   "Carrier_81_G120DStatusWord.9" AT %I4413.1 : Bool;   // Bit_09_CONTR_PLC
   "Carrier_81_G120DStatusWord.10" AT %I4413.2 : Bool;   // Bit_10_F_MAX
   "Carrier_81_G120DStatusWord.11" AT %I4413.3 : Bool;   // Bit_11_LIMIT_REACHED
   "Carrier_81_G120DStatusWord.12" AT %I4413.4 : Bool;   // Bit_12_BRAKE_OPEN
   "Carrier_81_G120DStatusWord.13" AT %I4413.5 : Bool;   // Bit_13_NO_OVERTEMP
   "Carrier_81_G120DStatusWord.14" AT %I4413.6 : Bool;   // Bit_14_CW_CCW
   "Carrier_81_G120DStatusWord.15" AT %I4413.7 : Bool;   // Bit_15_OVERL
   "Carrier_81_Slot2_Input" AT %IW4414 : Word;   // SLOT 2 INPUT WORD
   "Carrier_81_CrashDetectSW" AT %I4414.0 : Bool;   // CRASH DETECT SW
   "Carrier_81_SpareSafetyInput(2_1)" AT %I4414.1 : Bool;   // SPARE SAFETY INPUT
   "Carrier_81_SpareSafetyInput(2_2)" AT %I4414.2 : Bool;   // SPARE SAFETY INPUT
   "Carrier_81_SpareSafetyInput(2_3)" AT %I4414.3 : Bool;   // SPARE SAFETY INPUT
   "Carrier_81_SpareSafetyInput(2_4)" AT %I4414.4 : Bool;   // SPARE SAFETY INPUT
   "Carrier_81_SpareSafetyInput(2_5)" AT %I4414.5 : Bool;   // SPARE SAFETY INPUT
   "Carrier_81_SpareSafetyInput(2_6)" AT %I4414.6 : Bool;   // SPARE SAFETY INPUT
   "Carrier_81_SpareSafetyInput(2_7)" AT %I4414.7 : Bool;   // SPARE SAFETY INPUT
   "Carrier_81_Slot3_SafetyOutput" AT %IW4415 : Word;   // SLOT 3 SAFETY OUTPUT WORD
   "Carrier_81_Crash_Detect_OK" AT %I4415.0 : Bool;   // CARRIER CRASH DETECT
   "Carrier_81_SpareSafetyOutput(3_1)" AT %I4415.1 : Bool;   // SPARE SAFETY OUTPUT
   "Carrier_81_SpareSafetyOutput(3_2)" AT %I4415.2 : Bool;   // SPARE SAFETY OUTPUT
   "Carrier_81_SpareSafetyOutput(3_3)" AT %I4415.3 : Bool;   // SPARE SAFETY OUTPUT
   "Carrier_81_SpareSafetyOutput(3_4)" AT %I4415.4 : Bool;   // SPARE SAFETY OUTPUT
   "Carrier_81_SpareSafetyOutput(3_5)" AT %I4415.5 : Bool;   // SPARE SAFETY OUTPUT
   "Carrier_81_SpareSafetyOutput(3_6)" AT %I4415.6 : Bool;   // SPARE SAFETY OUTPUT
   "Carrier_81_SpareSafetyOutput(3_7)" AT %I4415.7 : Bool;   // SPARE SAFETY OUTPUT
   "Carrier_81_Slot4_Input" AT %IW4416 : Word;   // SLOT 4 INPUT WORD
   "Carrier_81_480VPowerOn_MDCB1" AT %I4416.0 : Bool;   // 480 VAC POWER ON MDCB 1
   "Carrier_81_SpareInput(4_1)" AT %I4416.1 : Bool;   // SPARE INPUT
   "Carrier_81_SpareInput(4_2)" AT %I4416.2 : Bool;   // SPARE INPUT
   "Carrier_81_SitopSelectStatus" AT %I4416.3 : Bool;   // SITOP SELECT STATUS
   "Carrier_81_DCsupplyOnPSCB2" AT %I4416.4 : Bool;   // DC SUPPLY ON PSCB 2
   "Carrier_81_SpareInput(4_5)" AT %I4416.5 : Bool;   // SPARE INPUT
   "Carrier_81_SpareInput(4_6)" AT %I4416.6 : Bool;   // SPARE INPUT
   "Carrier_81_SpareInput(4_7)" AT %I4416.7 : Bool;   // SPARE INPUT
   "Carrier_81_PB1_ProdHoldLH" AT %I4417.0 : Bool;   // PB 1 PRODUCTION HOLD LH
   "Carrier_81_PB2_ResetLH" AT %I4417.1 : Bool;   // PB 2 RESET LH
   "Carrier_81_PB3_ProdHoldRH" AT %I4417.2 : Bool;   // PB 3 PRODUCTION HOLD RH
   "Carrier_81_PB4_ResetRH" AT %I4417.3 : Bool;   // PB 4 RESET RH
   "Carrier_81_SpareInput(4_14)" AT %I4417.4 : Bool;   // SPARE INPUT
   "Carrier_81_SpareInput(4_15)" AT %I4417.5 : Bool;   // SPARE INPUT
   "Carrier_81_SpareInput(4_16)" AT %I4417.6 : Bool;   // SPARE INPUT
   "Carrier_81_SpareInput(4_17)" AT %I4417.7 : Bool;   // SPARE INPUT
   "Carrier_81_Slot5_Output" AT %IW4418 : Word;   // SLOT 5 OUTPUT WORD
   "Carrier_81_IRD400_HMI_24VDC_ENABLE" AT %I4418.0 : Bool;   // IRD 400 PANEL HMI 24V DC POWER
   "Carrier_81_FaultLight_LH" AT %I4418.1 : Bool;   // FAULT LIGHT LH
   "Carrier_81_RunLight_LH" AT %I4418.2 : Bool;   // RUN LIGHT LH
   "Carrier_81_FaultLight_RH" AT %I4418.3 : Bool;   // FAULT LIGHT RH
   "Carrier_81_RunLight_RH" AT %I4418.4 : Bool;   // RUN LIGHT RH
   "Carrier_81_SpareOutput(5_5)" AT %I4418.5 : Bool;   // SPARE OUTPUT
   "Carrier_81_SpareOutput(5_6)" AT %I4418.6 : Bool;   // SPARE OUTPUT
   "Carrier_81_SpareOutput(5_7)" AT %I4418.7 : Bool;   // SPARE OUTPUT
   "Carrier_81_ActualSpeed" AT %IW4420 : Word;   // ACTUAL SPEED
   "Carrier_81_CarrierDriveAlarm" AT %IW4422 : Word;   // CARRIER DRIVE ALARM
   "Carrier_81_CarrierDriveWarning" AT %IW4424 : Word;   // CARRIER DRIVE WARNING
   "Carrier_82_Status" AT %IW4450 : Word;   // CARRIER STATUS WORD
   "Carrier_82_Status.0" AT %I4450.0 : Bool;   // HEARTBEAT
   "Carrier_82_Status.1" AT %I4450.1 : Bool;   // MANUAL
   "Carrier_82_Status.2" AT %I4450.2 : Bool;   // IN_AUTO
   "Carrier_82_Status.3" AT %I4450.3 : Bool;   // POSITIONING_COMPLETE
   "Carrier_82_Status.4" AT %I4450.4 : Bool;   // PRODUCTION HOLD
   "Carrier_82_Status.5" AT %I4450.5 : Bool;   // CARRIER MOVING FORWARD
   "Carrier_82_Status.6" AT %I4450.6 : Bool;   // CARRIER MOVING REVERSE
   "Carrier_82_Status.7" AT %I4450.7 : Bool;   // CARRIER FAULT
   "Carrier_82_Status.8" AT %I4451.0 : Bool;   // CRASH DETECT TRIPPED
   "Carrier_82_Status.9" AT %I4451.1 : Bool;
   "Carrier_82_Status.10" AT %I4451.2 : Bool;
   "Carrier_82_Status.11" AT %I4451.3 : Bool;
   "Carrier_82_Status.12" AT %I4451.4 : Bool;
   "Carrier_82_Status.13" AT %I4451.5 : Bool;
   "Carrier_82_Status.14" AT %I4451.6 : Bool;
   "Carrier_82_Status.15" AT %I4451.7 : Bool;
   "Carrier_82_SDCFaultCode" AT %IW4452 : Word;   // SDC FAULT CODE
   "Carrier_82_CarrierPosition" AT %ID4454 : DWord;   // CARRIER POSITION
   "Carrier_82_CarrierNumber" AT %IW4458 : Word;   // CARRIER NUMBER
   "Carrier_82_G120DControlWord" AT %IW4460 : Word;   // G120D_STW1_CONTROL
   "Carrier_82_G120DControlWord.0" AT %I4460.0 : Bool;   // Bit_00_ON
   "Carrier_82_G120DControlWord.1" AT %I4460.1 : Bool;   // Bit_01_AUS2_INH
   "Carrier_82_G120DControlWord.2" AT %I4460.2 : Bool;   // Bit_02_AUS3_STOP
   "Carrier_82_G120DControlWord.3" AT %I4460.3 : Bool;   // Bit_03_EN
   "Carrier_82_G120DControlWord.4" AT %I4460.4 : Bool;   // Bit_04_EN_RAMP
   "Carrier_82_G120DControlWord.5" AT %I4460.5 : Bool;   // Bit_05_START_RAMP
   "Carrier_82_G120DControlWord.6" AT %I4460.6 : Bool;   // Bit_06_SETPOINT
   "Carrier_82_G120DControlWord.7" AT %I4460.7 : Bool;   // Bit_07_RESET
   "Carrier_82_G120DControlWord.8" AT %I4461.0 : Bool;   // Bit_08_JOG_R
   "Carrier_82_G120DControlWord.9" AT %I4461.1 : Bool;   // Bit_09_JOG_L
   "Carrier_82_G120DControlWord.10" AT %I4461.2 : Bool;   // Bit_10_CONTR_PLC
   "Carrier_82_G120DControlWord.11" AT %I4461.3 : Bool;   // Bit_11_REVERSE
   "Carrier_82_G120DControlWord.12" AT %I4461.4 : Bool;   // Bit_12_BRAKE_RELEASE
   "Carrier_82_G120DControlWord.13" AT %I4461.5 : Bool;   // Bit_13_DDS
   "Carrier_82_G120DControlWord.14" AT %I4461.6 : Bool;   // Bit_14_DO0
   "Carrier_82_G120DControlWord.15" AT %I4461.7 : Bool;   // Bit_15_DO1
   "Carrier_82_G120DStatusWord" AT %IW4462 : Word;   // G120D_ZSW1_STATUS
   "Carrier_82_G120DStatusWord.0" AT %I4462.0 : Bool;   // Bit_00_READY_RUN
   "Carrier_82_G120DStatusWord.1" AT %I4462.1 : Bool;   // Bit_01_READY_ON
   "Carrier_82_G120DStatusWord.2" AT %I4462.2 : Bool;   // Bit_02_ENABLE
   "Carrier_82_G120DStatusWord.3" AT %I4462.3 : Bool;   // Bit_03_FAULT
   "Carrier_82_G120DStatusWord.4" AT %I4462.4 : Bool;   // Bit_04_OFF2
   "Carrier_82_G120DStatusWord.5" AT %I4462.5 : Bool;   // Bit_05_OFF3
   "Carrier_82_G120DStatusWord.6" AT %I4462.6 : Bool;   // Bit_06_LOCK_OUT
   "Carrier_82_G120DStatusWord.7" AT %I4462.7 : Bool;   // Bit_07_WARN
   "Carrier_82_G120DStatusWord.8" AT %I4463.0 : Bool;   // Bit_08_NO_DEVIATION
   "Carrier_82_G120DStatusWord.9" AT %I4463.1 : Bool;   // Bit_09_CONTR_PLC
   "Carrier_82_G120DStatusWord.10" AT %I4463.2 : Bool;   // Bit_10_F_MAX
   "Carrier_82_G120DStatusWord.11" AT %I4463.3 : Bool;   // Bit_11_LIMIT_REACHED
   "Carrier_82_G120DStatusWord.12" AT %I4463.4 : Bool;   // Bit_12_BRAKE_OPEN
   "Carrier_82_G120DStatusWord.13" AT %I4463.5 : Bool;   // Bit_13_NO_OVERTEMP
   "Carrier_82_G120DStatusWord.14" AT %I4463.6 : Bool;   // Bit_14_CW_CCW
   "Carrier_82_G120DStatusWord.15" AT %I4463.7 : Bool;   // Bit_15_OVERL
   "Carrier_82_Slot2_Input" AT %IW4464 : Word;   // SLOT 2 INPUT WORD
   "Carrier_82_CrashDetectSW" AT %I4464.0 : Bool;   // CRASH DETECT SW
   "Carrier_82_SpareSafetyInput(2_1)" AT %I4464.1 : Bool;   // SPARE SAFETY INPUT
   "Carrier_82_SpareSafetyInput(2_2)" AT %I4464.2 : Bool;   // SPARE SAFETY INPUT
   "Carrier_82_SpareSafetyInput(2_3)" AT %I4464.3 : Bool;   // SPARE SAFETY INPUT
   "Carrier_82_SpareSafetyInput(2_4)" AT %I4464.4 : Bool;   // SPARE SAFETY INPUT
   "Carrier_82_SpareSafetyInput(2_5)" AT %I4464.5 : Bool;   // SPARE SAFETY INPUT
   "Carrier_82_SpareSafetyInput(2_6)" AT %I4464.6 : Bool;   // SPARE SAFETY INPUT
   "Carrier_82_SpareSafetyInput(2_7)" AT %I4464.7 : Bool;   // SPARE SAFETY INPUT
   "Carrier_82_Slot3_SafetyOutput" AT %IW4465 : Word;   // SLOT 3 SAFETY OUTPUT WORD
   "Carrier_82_Crash_Detect_OK" AT %I4465.0 : Bool;   // CARRIER CRASH DETECT
   "Carrier_82_SpareSafetyOutput(3_1)" AT %I4465.1 : Bool;   // SPARE SAFETY OUTPUT
   "Carrier_82_SpareSafetyOutput(3_2)" AT %I4465.2 : Bool;   // SPARE SAFETY OUTPUT
   "Carrier_82_SpareSafetyOutput(3_3)" AT %I4465.3 : Bool;   // SPARE SAFETY OUTPUT
   "Carrier_82_SpareSafetyOutput(3_4)" AT %I4465.4 : Bool;   // SPARE SAFETY OUTPUT
   "Carrier_82_SpareSafetyOutput(3_5)" AT %I4465.5 : Bool;   // SPARE SAFETY OUTPUT
   "Carrier_82_SpareSafetyOutput(3_6)" AT %I4465.6 : Bool;   // SPARE SAFETY OUTPUT
   "Carrier_82_SpareSafetyOutput(3_7)" AT %I4465.7 : Bool;   // SPARE SAFETY OUTPUT
   "Carrier_82_Slot4_Input" AT %IW4466 : Word;   // SLOT 4 INPUT WORD
   "Carrier_82_480VPowerOn_MDCB1" AT %I4466.0 : Bool;   // 480 VAC POWER ON MDCB 1
   "Carrier_82_SpareInput(4_1)" AT %I4466.1 : Bool;   // SPARE INPUT
   "Carrier_82_SpareInput(4_2)" AT %I4466.2 : Bool;   // SPARE INPUT
   "Carrier_82_SitopSelectStatus" AT %I4466.3 : Bool;   // SITOP SELECT STATUS
   "Carrier_82_DCsupplyOnPSCB2" AT %I4466.4 : Bool;   // DC SUPPLY ON PSCB 2
   "Carrier_82_SpareInput(4_5)" AT %I4466.5 : Bool;   // SPARE INPUT
   "Carrier_82_SpareInput(4_6)" AT %I4466.6 : Bool;   // SPARE INPUT
   "Carrier_82_SpareInput(4_7)" AT %I4466.7 : Bool;   // SPARE INPUT
   "Carrier_82_PB1_ProdHoldLH" AT %I4467.0 : Bool;   // PB 1 PRODUCTION HOLD LH
   "Carrier_82_PB2_ResetLH" AT %I4467.1 : Bool;   // PB 2 RESET LH
   "Carrier_82_PB3_ProdHoldRH" AT %I4467.2 : Bool;   // PB 3 PRODUCTION HOLD RH
   "Carrier_82_PB4_ResetRH" AT %I4467.3 : Bool;   // PB 4 RESET RH
   "Carrier_82_SpareInput(4_14)" AT %I4467.4 : Bool;   // SPARE INPUT
   "Carrier_82_SpareInput(4_15)" AT %I4467.5 : Bool;   // SPARE INPUT
   "Carrier_82_SpareInput(4_16)" AT %I4467.6 : Bool;   // SPARE INPUT
   "Carrier_82_SpareInput(4_17)" AT %I4467.7 : Bool;   // SPARE INPUT
   "Carrier_82_Slot5_Output" AT %IW4468 : Word;   // SLOT 5 OUTPUT WORD
   "Carrier_82_IRD400_HMI_24VDC_ENABLE" AT %I4468.0 : Bool;   // IRD 400 PANEL HMI 24V DC POWER
   "Carrier_82_FaultLight_LH" AT %I4468.1 : Bool;   // FAULT LIGHT LH
   "Carrier_82_RunLight_LH" AT %I4468.2 : Bool;   // RUN LIGHT LH
   "Carrier_82_FaultLight_RH" AT %I4468.3 : Bool;   // FAULT LIGHT RH
   "Carrier_82_RunLight_RH" AT %I4468.4 : Bool;   // RUN LIGHT RH
   "Carrier_82_SpareOutput(5_5)" AT %I4468.5 : Bool;   // SPARE OUTPUT
   "Carrier_82_SpareOutput(5_6)" AT %I4468.6 : Bool;   // SPARE OUTPUT
   "Carrier_82_SpareOutput(5_7)" AT %I4468.7 : Bool;   // SPARE OUTPUT
   "Carrier_82_ActualSpeed" AT %IW4470 : Word;   // ACTUAL SPEED
   "Carrier_82_CarrierDriveAlarm" AT %IW4472 : Word;   // CARRIER DRIVE ALARM
   "Carrier_82_CarrierDriveWarning" AT %IW4474 : Word;   // CARRIER DRIVE WARNING
   "Tag_101" AT %M2.3 : Bool;
   "Tag_100" AT %M3.7 : Bool;
   "Tag_117" AT %MW58 : Word;
END_VAR

VAR_GLOBAL   // PLC tag table "SDC_Carrier_TagTable"
   "Carrier_01_Carrier_In_Zone" AT %QW400 : Word;
   "Carrier_01_Carrier_Number_Echo" AT %QW402 : Word;
   "Carrier_01_Carrier_Position_Echo" AT %QD404 : DWord;
   "Carrier_01_Next_Carrier_Number" AT %QW408 : Word;
   "Carrier_01_Next_Stop_Position" AT %QD410 : DWord;
   "Carrier_01_Drive_Command_Speed" AT %QW414 : Word;
   "Carrier_01_Duplicate_Carrier_Number" AT %QW416 : Word;
   "Carrier_01_First_Duplicate_Carrier_Position" AT %QD418 : DWord;
   "Carrier_01_Second_Duplicate_Carrier_Position" AT %QD422 : DWord;
   "Carrier_01_CommandWord" AT %QW426 : Word;
   "Carrier_01_Heartbeat" AT %Q426.0 : Bool;
   "Carrier_01_Drive_Forward_Command" AT %Q426.1 : Bool;
   "Carrier_01_Fault_Reset" AT %Q426.2 : Bool;
   "Carrier_01_At_Command_Position" AT %Q426.3 : Bool;
   "Carrier_01_Duplicate_Carrier_Fault" AT %Q426.4 : Bool;
   "Carrier_01_Motion_On_Fault" AT %Q426.5 : Bool;
   "Carrier_01_Motion_Off_Fault" AT %Q426.6 : Bool;
   "Carrier_01_Carrier_Spacing_Fault" AT %Q426.7 : Bool;
   "Carrier_02_Carrier_In_Zone" AT %QW450 : Word;
   "Carrier_02_Carrier_Number_Echo" AT %QW452 : Word;
   "Carrier_02_Carrier_Position_Echo" AT %QD454 : DWord;
   "Carrier_02_Next_Carrier_Number" AT %QW458 : Word;
   "Carrier_02_Next_Stop_Position" AT %QD460 : DWord;
   "Carrier_02_Drive_Command_Speed" AT %QW464 : Word;
   "Carrier_02_Duplicate_Carrier_Number" AT %QW466 : Word;
   "Carrier_02_First_Duplicate_Carrier_Position" AT %QD468 : DWord;
   "Carrier_02_Second_Duplicate_Carrier_Position" AT %QD472 : DWord;
   "Carrier_02_CommandWord" AT %QW476 : Word;
   "Carrier_02_Heartbeat" AT %Q476.0 : Bool;
   "Carrier_02_Drive_Forward_Command" AT %Q476.1 : Bool;
   "Carrier_02_Fault_Reset" AT %Q476.2 : Bool;
   "Carrier_02_At_Command_Position" AT %Q476.3 : Bool;
   "Carrier_02_Duplicate_Carrier_Fault" AT %Q476.4 : Bool;
   "Carrier_02_Motion_On_Fault" AT %Q476.5 : Bool;
   "Carrier_02_Motion_Off_Fault" AT %Q476.6 : Bool;
   "Carrier_02_Carrier_Spacing_Fault" AT %Q476.7 : Bool;
   "Carrier_03_Carrier_In_Zone" AT %QW500 : Word;
   "Carrier_03_Carrier_Number_Echo" AT %QW502 : Word;
   "Carrier_03_Carrier_Position_Echo" AT %QD504 : DWord;
   "Carrier_03_Next_Carrier_Number" AT %QW508 : Word;
   "Carrier_03_Next_Stop_Position" AT %QD510 : DWord;
   "Carrier_03_Drive_Command_Speed" AT %QW514 : Word;
   "Carrier_03_Duplicate_Carrier_Number" AT %QW516 : Word;
   "Carrier_03_First_Duplicate_Carrier_Position" AT %QD518 : DWord;
   "Carrier_03_Second_Duplicate_Carrier_Position" AT %QD522 : DWord;
   "Carrier_03_CommandWord" AT %QW526 : Word;
   "Carrier_03_Heartbeat" AT %Q526.0 : Bool;
   "Carrier_03_Drive_Forward_Command" AT %Q526.1 : Bool;
   "Carrier_03_Fault_Reset" AT %Q526.2 : Bool;
   "Carrier_03_At_Command_Position" AT %Q526.3 : Bool;
   "Carrier_03_Duplicate_Carrier_Fault" AT %Q526.4 : Bool;
   "Carrier_03_Motion_On_Fault" AT %Q526.5 : Bool;
   "Carrier_03_Motion_Off_Fault" AT %Q526.6 : Bool;
   "Carrier_03_Carrier_Spacing_Fault" AT %Q526.7 : Bool;
   "Carrier_04_Carrier_In_Zone" AT %QW550 : Word;
   "Carrier_04_Carrier_Number_Echo" AT %QW552 : Word;
   "Carrier_04_Carrier_Position_Echo" AT %QD554 : DWord;
   "Carrier_04_Next_Carrier_Number" AT %QW558 : Word;
   "Carrier_04_Next_Stop_Position" AT %QD560 : DWord;
   "Carrier_04_Drive_Command_Speed" AT %QW564 : Word;
   "Carrier_04_Duplicate_Carrier_Number" AT %QW566 : Word;
   "Carrier_04_First_Duplicate_Carrier_Position" AT %QD568 : DWord;
   "Carrier_04_Second_Duplicate_Carrier_Position" AT %QD572 : DWord;
   "Carrier_04_CommandWord" AT %QW576 : Word;
   "Carrier_04_Heartbeat" AT %Q576.0 : Bool;
   "Carrier_04_Drive_Forward_Command" AT %Q576.1 : Bool;
   "Carrier_04_Fault_Reset" AT %Q576.2 : Bool;
   "Carrier_04_At_Command_Position" AT %Q576.3 : Bool;
   "Carrier_04_Duplicate_Carrier_Fault" AT %Q576.4 : Bool;
   "Carrier_04_Motion_On_Fault" AT %Q576.5 : Bool;
   "Carrier_04_Motion_Off_Fault" AT %Q576.6 : Bool;
   "Carrier_04_Carrier_Spacing_Fault" AT %Q576.7 : Bool;
   "Carrier_05_Carrier_In_Zone" AT %QW600 : Word;
   "Carrier_05_Carrier_Number_Echo" AT %QW602 : Word;
   "Carrier_05_Carrier_Position_Echo" AT %QD604 : DWord;
   "Carrier_05_Next_Carrier_Number" AT %QW608 : Word;
   "Carrier_05_Next_Stop_Position" AT %QD610 : DWord;
   "Carrier_05_Drive_Command_Speed" AT %QW614 : Word;
   "Carrier_05_Duplicate_Carrier_Number" AT %QW616 : Word;
   "Carrier_05_First_Duplicate_Carrier_Position" AT %QD618 : DWord;
   "Carrier_05_Second_Duplicate_Carrier_Position" AT %QD622 : DWord;
   "Carrier_05_CommandWord" AT %QW626 : Word;
   "Carrier_05_Heartbeat" AT %Q626.0 : Bool;
   "Carrier_05_Drive_Forward_Command" AT %Q626.1 : Bool;
   "Carrier_05_Fault_Reset" AT %Q626.2 : Bool;
   "Carrier_05_At_Command_Position" AT %Q626.3 : Bool;
   "Carrier_05_Duplicate_Carrier_Fault" AT %Q626.4 : Bool;
   "Carrier_05_Motion_On_Fault" AT %Q626.5 : Bool;
   "Carrier_05_Motion_Off_Fault" AT %Q626.6 : Bool;
   "Carrier_05_Carrier_Spacing_Fault" AT %Q626.7 : Bool;
   "Carrier_06_Carrier_In_Zone" AT %QW650 : Word;
   "Carrier_06_Carrier_Number_Echo" AT %QW652 : Word;
   "Carrier_06_Carrier_Position_Echo" AT %QD654 : DWord;
   "Carrier_06_Next_Carrier_Number" AT %QW658 : Word;
   "Carrier_06_Next_Stop_Position" AT %QD660 : DWord;
   "Carrier_06_Drive_Command_Speed" AT %QW664 : Word;
   "Carrier_06_Duplicate_Carrier_Number" AT %QW666 : Word;
   "Carrier_06_First_Duplicate_Carrier_Position" AT %QD668 : DWord;
   "Carrier_06_Second_Duplicate_Carrier_Position" AT %QD672 : DWord;
   "Carrier_06_CommandWord" AT %QW676 : Word;
   "Carrier_06_Heartbeat" AT %Q676.0 : Bool;
   "Carrier_06_Drive_Forward_Command" AT %Q676.1 : Bool;
   "Carrier_06_Fault_Reset" AT %Q676.2 : Bool;
   "Carrier_06_At_Command_Position" AT %Q676.3 : Bool;
   "Carrier_06_Duplicate_Carrier_Fault" AT %Q676.4 : Bool;
   "Carrier_06_Motion_On_Fault" AT %Q676.5 : Bool;
   "Carrier_06_Motion_Off_Fault" AT %Q676.6 : Bool;
   "Carrier_06_Carrier_Spacing_Fault" AT %Q676.7 : Bool;
   "Carrier_07_Carrier_In_Zone" AT %QW700 : Word;
   "Carrier_07_Carrier_Number_Echo" AT %QW702 : Word;
   "Carrier_07_Carrier_Position_Echo" AT %QD704 : DWord;
   "Carrier_07_Next_Carrier_Number" AT %QW708 : Word;
   "Carrier_07_Next_Stop_Position" AT %QD710 : DWord;
   "Carrier_07_Drive_Command_Speed" AT %QW714 : Word;
   "Carrier_07_Duplicate_Carrier_Number" AT %QW716 : Word;
   "Carrier_07_First_Duplicate_Carrier_Position" AT %QD718 : DWord;
   "Carrier_07_Second_Duplicate_Carrier_Position" AT %QD722 : DWord;
   "Carrier_07_CommandWord" AT %QW726 : Word;
   "Carrier_07_Heartbeat" AT %Q726.0 : Bool;
   "Carrier_07_Drive_Forward_Command" AT %Q726.1 : Bool;
   "Carrier_07_Fault_Reset" AT %Q726.2 : Bool;
   "Carrier_07_At_Command_Position" AT %Q726.3 : Bool;
   "Carrier_07_Duplicate_Carrier_Fault" AT %Q726.4 : Bool;
   "Carrier_07_Motion_On_Fault" AT %Q726.5 : Bool;
   "Carrier_07_Motion_Off_Fault" AT %Q726.6 : Bool;
   "Carrier_07_Carrier_Spacing_Fault" AT %Q726.7 : Bool;
   "Carrier_08_Carrier_In_Zone" AT %QW750 : Word;
   "Carrier_08_Carrier_Number_Echo" AT %QW752 : Word;
   "Carrier_08_Carrier_Position_Echo" AT %QD754 : DWord;
   "Carrier_08_Next_Carrier_Number" AT %QW758 : Word;
   "Carrier_08_Next_Stop_Position" AT %QD760 : DWord;
   "Carrier_08_Drive_Command_Speed" AT %QW764 : Word;
   "Carrier_08_Duplicate_Carrier_Number" AT %QW766 : Word;
   "Carrier_08_First_Duplicate_Carrier_Position" AT %QD768 : DWord;
   "Carrier_08_Second_Duplicate_Carrier_Position" AT %QD772 : DWord;
   "Carrier_08_CommandWord" AT %QW776 : Word;
   "Carrier_08_Heartbeat" AT %Q776.0 : Bool;
   "Carrier_08_Drive_Forward_Command" AT %Q776.1 : Bool;
   "Carrier_08_Fault_Reset" AT %Q776.2 : Bool;
   "Carrier_08_At_Command_Position" AT %Q776.3 : Bool;
   "Carrier_08_Duplicate_Carrier_Fault" AT %Q776.4 : Bool;
   "Carrier_08_Motion_On_Fault" AT %Q776.5 : Bool;
   "Carrier_08_Motion_Off_Fault" AT %Q776.6 : Bool;
   "Carrier_08_Carrier_Spacing_Fault" AT %Q776.7 : Bool;
   "Carrier_09_Carrier_In_Zone" AT %QW800 : Word;
   "Carrier_09_Carrier_Number_Echo" AT %QW802 : Word;
   "Carrier_09_Carrier_Position_Echo" AT %QD804 : DWord;
   "Carrier_09_Next_Carrier_Number" AT %QW808 : Word;
   "Carrier_09_Next_Stop_Position" AT %QD810 : DWord;
   "Carrier_09_Drive_Command_Speed" AT %QW814 : Word;
   "Carrier_09_Duplicate_Carrier_Number" AT %QW816 : Word;
   "Carrier_09_First_Duplicate_Carrier_Position" AT %QD818 : DWord;
   "Carrier_09_Second_Duplicate_Carrier_Position" AT %QD822 : DWord;
   "Carrier_09_CommandWord" AT %QW826 : Word;
   "Carrier_09_Heartbeat" AT %Q826.0 : Bool;
   "Carrier_09_Drive_Forward_Command" AT %Q826.1 : Bool;
   "Carrier_09_Fault_Reset" AT %Q826.2 : Bool;
   "Carrier_09_At_Command_Position" AT %Q826.3 : Bool;
   "Carrier_09_Duplicate_Carrier_Fault" AT %Q826.4 : Bool;
   "Carrier_09_Motion_On_Fault" AT %Q826.5 : Bool;
   "Carrier_09_Motion_Off_Fault" AT %Q826.6 : Bool;
   "Carrier_09_Carrier_Spacing_Fault" AT %Q826.7 : Bool;
   "Carrier_10_Carrier_In_Zone" AT %QW850 : Word;
   "Carrier_10_Carrier_Number_Echo" AT %QW852 : Word;
   "Carrier_10_Carrier_Position_Echo" AT %QD854 : DWord;
   "Carrier_10_Next_Carrier_Number" AT %QW858 : Word;
   "Carrier_10_Next_Stop_Position" AT %QD860 : DWord;
   "Carrier_10_Drive_Command_Speed" AT %QW864 : Word;
   "Carrier_10_Duplicate_Carrier_Number" AT %QW866 : Word;
   "Carrier_10_First_Duplicate_Carrier_Position" AT %QD868 : DWord;
   "Carrier_10_Second_Duplicate_Carrier_Position" AT %QD872 : DWord;
   "Carrier_10_CommandWord" AT %QW876 : Word;
   "Carrier_10_Heartbeat" AT %Q876.0 : Bool;
   "Carrier_10_Drive_Forward_Command" AT %Q876.1 : Bool;
   "Carrier_10_Fault_Reset" AT %Q876.2 : Bool;
   "Carrier_10_At_Command_Position" AT %Q876.3 : Bool;
   "Carrier_10_Duplicate_Carrier_Fault" AT %Q876.4 : Bool;
   "Carrier_10_Motion_On_Fault" AT %Q876.5 : Bool;
   "Carrier_10_Motion_Off_Fault" AT %Q876.6 : Bool;
   "Carrier_10_Carrier_Spacing_Fault" AT %Q876.7 : Bool;
   "Carrier_11_Carrier_In_Zone" AT %QW900 : Word;
   "Carrier_11_Carrier_Number_Echo" AT %QW902 : Word;
   "Carrier_11_Carrier_Position_Echo" AT %QD904 : DWord;
   "Carrier_11_Next_Carrier_Number" AT %QW908 : Word;
   "Carrier_11_Next_Stop_Position" AT %QD910 : DWord;
   "Carrier_11_Drive_Command_Speed" AT %QW914 : Word;
   "Carrier_11_Duplicate_Carrier_Number" AT %QW916 : Word;
   "Carrier_11_First_Duplicate_Carrier_Position" AT %QD918 : DWord;
   "Carrier_11_Second_Duplicate_Carrier_Position" AT %QD922 : DWord;
   "Carrier_11_CommandWord" AT %QW926 : Word;
   "Carrier_11_Heartbeat" AT %Q926.0 : Bool;
   "Carrier_11_Drive_Forward_Command" AT %Q926.1 : Bool;
   "Carrier_11_Fault_Reset" AT %Q926.2 : Bool;
   "Carrier_11_At_Command_Position" AT %Q926.3 : Bool;
   "Carrier_11_Duplicate_Carrier_Fault" AT %Q926.4 : Bool;
   "Carrier_11_Motion_On_Fault" AT %Q926.5 : Bool;
   "Carrier_11_Motion_Off_Fault" AT %Q926.6 : Bool;
   "Carrier_11_Carrier_Spacing_Fault" AT %Q926.7 : Bool;
   "Carrier_12_Carrier_In_Zone" AT %QW950 : Word;
   "Carrier_12_Carrier_Number_Echo" AT %QW952 : Word;
   "Carrier_12_Carrier_Position_Echo" AT %QD954 : DWord;
   "Carrier_12_Next_Carrier_Number" AT %QW958 : Word;
   "Carrier_12_Next_Stop_Position" AT %QD960 : DWord;
   "Carrier_12_Drive_Command_Speed" AT %QW964 : Word;
   "Carrier_12_Duplicate_Carrier_Number" AT %QW966 : Word;
   "Carrier_12_First_Duplicate_Carrier_Position" AT %QD968 : DWord;
   "Carrier_12_Second_Duplicate_Carrier_Position" AT %QD972 : DWord;
   "Carrier_12_CommandWord" AT %QW976 : Word;
   "Carrier_12_Heartbeat" AT %Q976.0 : Bool;
   "Carrier_12_Drive_Forward_Command" AT %Q976.1 : Bool;
   "Carrier_12_Fault_Reset" AT %Q976.2 : Bool;
   "Carrier_12_At_Command_Position" AT %Q976.3 : Bool;
   "Carrier_12_Duplicate_Carrier_Fault" AT %Q976.4 : Bool;
   "Carrier_12_Motion_On_Fault" AT %Q976.5 : Bool;
   "Carrier_12_Motion_Off_Fault" AT %Q976.6 : Bool;
   "Carrier_12_Carrier_Spacing_Fault" AT %Q976.7 : Bool;
   "Carrier_13_Carrier_In_Zone" AT %QW1000 : Word;
   "Carrier_13_Carrier_Number_Echo" AT %QW1002 : Word;
   "Carrier_13_Carrier_Position_Echo" AT %QD1004 : DWord;
   "Carrier_13_Next_Carrier_Number" AT %QW1008 : Word;
   "Carrier_13_Next_Stop_Position" AT %QD1010 : DWord;
   "Carrier_13_Drive_Command_Speed" AT %QW1014 : Word;
   "Carrier_13_Duplicate_Carrier_Number" AT %QW1016 : Word;
   "Carrier_13_First_Duplicate_Carrier_Position" AT %QD1018 : DWord;
   "Carrier_13_Second_Duplicate_Carrier_Position" AT %QD1022 : DWord;
   "Carrier_13_CommandWord" AT %QW1026 : Word;
   "Carrier_13_Heartbeat" AT %Q1026.0 : Bool;
   "Carrier_13_Drive_Forward_Command" AT %Q1026.1 : Bool;
   "Carrier_13_Fault_Reset" AT %Q1026.2 : Bool;
   "Carrier_13_At_Command_Position" AT %Q1026.3 : Bool;
   "Carrier_13_Duplicate_Carrier_Fault" AT %Q1026.4 : Bool;
   "Carrier_13_Motion_On_Fault" AT %Q1026.5 : Bool;
   "Carrier_13_Motion_Off_Fault" AT %Q1026.6 : Bool;
   "Carrier_13_Carrier_Spacing_Fault" AT %Q1026.7 : Bool;
   "Carrier_14_Carrier_In_Zone" AT %QW1050 : Word;
   "Carrier_14_Carrier_Number_Echo" AT %QW1052 : Word;
   "Carrier_14_Carrier_Position_Echo" AT %QD1054 : DWord;
   "Carrier_14_Next_Carrier_Number" AT %QW1058 : Word;
   "Carrier_14_Next_Stop_Position" AT %QD1060 : DWord;
   "Carrier_14_Drive_Command_Speed" AT %QW1064 : Word;
   "Carrier_14_Duplicate_Carrier_Number" AT %QW1066 : Word;
   "Carrier_14_First_Duplicate_Carrier_Position" AT %QD1068 : DWord;
   "Carrier_14_Second_Duplicate_Carrier_Position" AT %QD1072 : DWord;
   "Carrier_14_CommandWord" AT %QW1076 : Word;
   "Carrier_14_Heartbeat" AT %Q1076.0 : Bool;
   "Carrier_14_Drive_Forward_Command" AT %Q1076.1 : Bool;
   "Carrier_14_Fault_Reset" AT %Q1076.2 : Bool;
   "Carrier_14_At_Command_Position" AT %Q1076.3 : Bool;
   "Carrier_14_Duplicate_Carrier_Fault" AT %Q1076.4 : Bool;
   "Carrier_14_Motion_On_Fault" AT %Q1076.5 : Bool;
   "Carrier_14_Motion_Off_Fault" AT %Q1076.6 : Bool;
   "Carrier_14_Carrier_Spacing_Fault" AT %Q1076.7 : Bool;
   "Carrier_15_Carrier_In_Zone" AT %QW1100 : Word;
   "Carrier_15_Carrier_Number_Echo" AT %QW1102 : Word;
   "Carrier_15_Carrier_Position_Echo" AT %QD1104 : DWord;
   "Carrier_15_Next_Carrier_Number" AT %QW1108 : Word;
   "Carrier_15_Next_Stop_Position" AT %QD1110 : DWord;
   "Carrier_15_Drive_Command_Speed" AT %QW1114 : Word;
   "Carrier_15_Duplicate_Carrier_Number" AT %QW1116 : Word;
   "Carrier_15_First_Duplicate_Carrier_Position" AT %QD1118 : DWord;
   "Carrier_15_Second_Duplicate_Carrier_Position" AT %QD1122 : DWord;
   "Carrier_15_CommandWord" AT %QW1126 : Word;
   "Carrier_15_Heartbeat" AT %Q1126.0 : Bool;
   "Carrier_15_Drive_Forward_Command" AT %Q1126.1 : Bool;
   "Carrier_15_Fault_Reset" AT %Q1126.2 : Bool;
   "Carrier_15_At_Command_Position" AT %Q1126.3 : Bool;
   "Carrier_15_Duplicate_Carrier_Fault" AT %Q1126.4 : Bool;
   "Carrier_15_Motion_On_Fault" AT %Q1126.5 : Bool;
   "Carrier_15_Motion_Off_Fault" AT %Q1126.6 : Bool;
   "Carrier_15_Carrier_Spacing_Fault" AT %Q1126.7 : Bool;
   "Carrier_16_Carrier_In_Zone" AT %QW1150 : Word;
   "Carrier_16_Carrier_Number_Echo" AT %QW1152 : Word;
   "Carrier_16_Carrier_Position_Echo" AT %QD1154 : DWord;
   "Carrier_16_Next_Carrier_Number" AT %QW1158 : Word;
   "Carrier_16_Next_Stop_Position" AT %QD1160 : DWord;
   "Carrier_16_Drive_Command_Speed" AT %QW1164 : Word;
   "Carrier_16_Duplicate_Carrier_Number" AT %QW1166 : Word;
   "Carrier_16_First_Duplicate_Carrier_Position" AT %QD1168 : DWord;
   "Carrier_16_Second_Duplicate_Carrier_Position" AT %QD1172 : DWord;
   "Carrier_16_CommandWord" AT %QW1176 : Word;
   "Carrier_16_Heartbeat" AT %Q1176.0 : Bool;
   "Carrier_16_Drive_Forward_Command" AT %Q1176.1 : Bool;
   "Carrier_16_Fault_Reset" AT %Q1176.2 : Bool;
   "Carrier_16_At_Command_Position" AT %Q1176.3 : Bool;
   "Carrier_16_Duplicate_Carrier_Fault" AT %Q1176.4 : Bool;
   "Carrier_16_Motion_On_Fault" AT %Q1176.5 : Bool;
   "Carrier_16_Motion_Off_Fault" AT %Q1176.6 : Bool;
   "Carrier_16_Carrier_Spacing_Fault" AT %Q1176.7 : Bool;
   "Carrier_17_Carrier_In_Zone" AT %QW1200 : Word;
   "Carrier_17_Carrier_Number_Echo" AT %QW1202 : Word;
   "Carrier_17_Carrier_Position_Echo" AT %QD1204 : DWord;
   "Carrier_17_Next_Carrier_Number" AT %QW1208 : Word;
   "Carrier_17_Next_Stop_Position" AT %QD1210 : DWord;
   "Carrier_17_Drive_Command_Speed" AT %QW1214 : Word;
   "Carrier_17_Duplicate_Carrier_Number" AT %QW1216 : Word;
   "Carrier_17_First_Duplicate_Carrier_Position" AT %QD1218 : DWord;
   "Carrier_17_Second_Duplicate_Carrier_Position" AT %QD1222 : DWord;
   "Carrier_17_CommandWord" AT %QW1226 : Word;
   "Carrier_17_Heartbeat" AT %Q1226.0 : Bool;
   "Carrier_17_Drive_Forward_Command" AT %Q1226.1 : Bool;
   "Carrier_17_Fault_Reset" AT %Q1226.2 : Bool;
   "Carrier_17_At_Command_Position" AT %Q1226.3 : Bool;
   "Carrier_17_Duplicate_Carrier_Fault" AT %Q1226.4 : Bool;
   "Carrier_17_Motion_On_Fault" AT %Q1226.5 : Bool;
   "Carrier_17_Motion_Off_Fault" AT %Q1226.6 : Bool;
   "Carrier_17_Carrier_Spacing_Fault" AT %Q1226.7 : Bool;
   "Carrier_18_Carrier_In_Zone" AT %QW1250 : Word;
   "Carrier_18_Carrier_Number_Echo" AT %QW1252 : Word;
   "Carrier_18_Carrier_Position_Echo" AT %QD1254 : DWord;
   "Carrier_18_Next_Carrier_Number" AT %QW1258 : Word;
   "Carrier_18_Next_Stop_Position" AT %QD1260 : DWord;
   "Carrier_18_Drive_Command_Speed" AT %QW1264 : Word;
   "Carrier_18_Duplicate_Carrier_Number" AT %QW1266 : Word;
   "Carrier_18_First_Duplicate_Carrier_Position" AT %QD1268 : DWord;
   "Carrier_18_Second_Duplicate_Carrier_Position" AT %QD1272 : DWord;
   "Carrier_18_CommandWord" AT %QW1276 : Word;
   "Carrier_18_Heartbeat" AT %Q1276.0 : Bool;
   "Carrier_18_Drive_Forward_Command" AT %Q1276.1 : Bool;
   "Carrier_18_Fault_Reset" AT %Q1276.2 : Bool;
   "Carrier_18_At_Command_Position" AT %Q1276.3 : Bool;
   "Carrier_18_Duplicate_Carrier_Fault" AT %Q1276.4 : Bool;
   "Carrier_18_Motion_On_Fault" AT %Q1276.5 : Bool;
   "Carrier_18_Motion_Off_Fault" AT %Q1276.6 : Bool;
   "Carrier_18_Carrier_Spacing_Fault" AT %Q1276.7 : Bool;
   "Carrier_19_Carrier_In_Zone" AT %QW1300 : Word;
   "Carrier_19_Carrier_Number_Echo" AT %QW1302 : Word;
   "Carrier_19_Carrier_Position_Echo" AT %QD1304 : DWord;
   "Carrier_19_Next_Carrier_Number" AT %QW1308 : Word;
   "Carrier_19_Next_Stop_Position" AT %QD1310 : DWord;
   "Carrier_19_Drive_Command_Speed" AT %QW1314 : Word;
   "Carrier_19_Duplicate_Carrier_Number" AT %QW1316 : Word;
   "Carrier_19_First_Duplicate_Carrier_Position" AT %QD1318 : DWord;
   "Carrier_19_Second_Duplicate_Carrier_Position" AT %QD1322 : DWord;
   "Carrier_19_CommandWord" AT %QW1326 : Word;
   "Carrier_19_Heartbeat" AT %Q1326.0 : Bool;
   "Carrier_19_Drive_Forward_Command" AT %Q1326.1 : Bool;
   "Carrier_19_Fault_Reset" AT %Q1326.2 : Bool;
   "Carrier_19_At_Command_Position" AT %Q1326.3 : Bool;
   "Carrier_19_Duplicate_Carrier_Fault" AT %Q1326.4 : Bool;
   "Carrier_19_Motion_On_Fault" AT %Q1326.5 : Bool;
   "Carrier_19_Motion_Off_Fault" AT %Q1326.6 : Bool;
   "Carrier_19_Carrier_Spacing_Fault" AT %Q1326.7 : Bool;
   "Carrier_20_Carrier_In_Zone" AT %QW1350 : Word;
   "Carrier_20_Carrier_Number_Echo" AT %QW1352 : Word;
   "Carrier_20_Carrier_Position_Echo" AT %QD1354 : DWord;
   "Carrier_20_Next_Carrier_Number" AT %QW1358 : Word;
   "Carrier_20_Next_Stop_Position" AT %QD1360 : DWord;
   "Carrier_20_Drive_Command_Speed" AT %QW1364 : Word;
   "Carrier_20_Duplicate_Carrier_Number" AT %QW1366 : Word;
   "Carrier_20_First_Duplicate_Carrier_Position" AT %QD1368 : DWord;
   "Carrier_20_Second_Duplicate_Carrier_Position" AT %QD1372 : DWord;
   "Carrier_20_CommandWord" AT %QW1376 : Word;
   "Carrier_20_Heartbeat" AT %Q1376.0 : Bool;
   "Carrier_20_Drive_Forward_Command" AT %Q1376.1 : Bool;
   "Carrier_20_Fault_Reset" AT %Q1376.2 : Bool;
   "Carrier_20_At_Command_Position" AT %Q1376.3 : Bool;
   "Carrier_20_Duplicate_Carrier_Fault" AT %Q1376.4 : Bool;
   "Carrier_20_Motion_On_Fault" AT %Q1376.5 : Bool;
   "Carrier_20_Motion_Off_Fault" AT %Q1376.6 : Bool;
   "Carrier_20_Carrier_Spacing_Fault" AT %Q1376.7 : Bool;
   "Carrier_21_Carrier_In_Zone" AT %QW1400 : Word;
   "Carrier_21_Carrier_Number_Echo" AT %QW1402 : Word;
   "Carrier_21_Carrier_Position_Echo" AT %QD1404 : DWord;
   "Carrier_21_Next_Carrier_Number" AT %QW1408 : Word;
   "Carrier_21_Next_Stop_Position" AT %QD1410 : DWord;
   "Carrier_21_Drive_Command_Speed" AT %QW1414 : Word;
   "Carrier_21_Duplicate_Carrier_Number" AT %QW1416 : Word;
   "Carrier_21_First_Duplicate_Carrier_Position" AT %QD1418 : DWord;
   "Carrier_21_Second_Duplicate_Carrier_Position" AT %QD1422 : DWord;
   "Carrier_21_CommandWord" AT %QW1426 : Word;
   "Carrier_21_Heartbeat" AT %Q1426.0 : Bool;
   "Carrier_21_Drive_Forward_Command" AT %Q1426.1 : Bool;
   "Carrier_21_Fault_Reset" AT %Q1426.2 : Bool;
   "Carrier_21_At_Command_Position" AT %Q1426.3 : Bool;
   "Carrier_21_Duplicate_Carrier_Fault" AT %Q1426.4 : Bool;
   "Carrier_21_Motion_On_Fault" AT %Q1426.5 : Bool;
   "Carrier_21_Motion_Off_Fault" AT %Q1426.6 : Bool;
   "Carrier_21_Carrier_Spacing_Fault" AT %Q1426.7 : Bool;
   "Carrier_22_Carrier_In_Zone" AT %QW1450 : Word;
   "Carrier_22_Carrier_Number_Echo" AT %QW1452 : Word;
   "Carrier_22_Carrier_Position_Echo" AT %QD1454 : DWord;
   "Carrier_22_Next_Carrier_Number" AT %QW1458 : Word;
   "Carrier_22_Next_Stop_Position" AT %QD1460 : DWord;
   "Carrier_22_Drive_Command_Speed" AT %QW1464 : Word;
   "Carrier_22_Duplicate_Carrier_Number" AT %QW1466 : Word;